DATA_BLOCK "PanelCompBAJA MTA"   // DB74
{ S7_Optimized_Access := 'FALSE' }
VERSION : 0.1
   VAR
      InhMC060 : Bool;
      InhMC061 : Bool;
      InhMC062 : Bool;
      InhMC063 : Bool;
      InhMC064 : Bool;
      InhMC065 : Bool;
      Flanco1MC060 : Bool;
      Flanco1MC061 : Bool;
      Flanco1MC062 : Bool;
      Flanco1MC063 : Bool;
      Flanco1MC064 : Bool;
      Flanco1MC065 : Bool;
      Flanco2MC060 : Bool;
      Flanco2MC061 : Bool;
      Flanco2MC062 : Bool;
      Flanco2MC063 : Bool;
      Flanco2MC064 : Bool;
      Flanco2MC065 : Bool;
      Flanco3MC060 : Bool;
      Flanco3MC061 : Bool;
      Flanco3MC062 : Bool;
      Flanco3MC063 : Bool;
      Flanco3MC064 : Bool;
      Flanco3MC065 : Bool;
      HabPanelMC060 : Bool;
      HabPanelMC061 : Bool;
      HabPanelMC062 : Bool;
      HabPanelMC063 : Bool;
      HabPanelMC064 : Bool;
      HabPanelMC065 : Bool;
      DeshabPanelMC060 : Bool;
      DeshabPanelMC061 : Bool;
      DeshabPanelMC062 : Bool;
      DeshabPanelMC063 : Bool;
      DeshabPanelMC064 : Bool;
      DeshabPanelMC065 : Bool;
      MarchaPanelMC060 : Bool;
      MarchaPanelMC061 : Bool;
      MarchaPanelMC062 : Bool;
      MarchaPanelMC063 : Bool;
      MarchaPanelMC064 : Bool;
      MarchaPanelMC065 : Bool;
      ParadaPanelMC060 : Bool;
      ParadaPanelMC061 : Bool;
      ParadaPanelMC062 : Bool;
      ParadaPanelMC063 : Bool;
      ParadaPanelMC064 : Bool;
      ParadaPanelMC065 : Bool;
      HabMC060 : Bool;
      HabMC061 : Bool;
      HabMC062 : Bool;
      HabMC063 : Bool;
      HabMC064 : Bool;
      HabMC065 : Bool;
      DeshabMC060 : Bool;
      DeshabMC061 : Bool;
      DeshabMC062 : Bool;
      DeshabMC063 : Bool;
      DeshabMC064 : Bool;
      DeshabMC065 : Bool;
      MarchaMC060 : Bool;
      MarchaMC061 : Bool;
      MarchaMC062 : Bool;
      MarchaMC063 : Bool;
      MarchaMC064 : Bool;
      MarchaMC065 : Bool;
      ParadaMC060 : Bool;
      ParadaMC061 : Bool;
      ParadaMC062 : Bool;
      ParadaMC063 : Bool;
      ParadaMC064 : Bool;
      ParadaMC065 : Bool;
      AnimMC060 : Byte;
      AnimMC061 : Byte;
      AnimMC062 : Byte;
      AnimMC063 : Byte;
      AnimMC064 : Byte;
      AnimMC065 : Byte;
      FallaGMTMC060 : Bool;
      FallaGMTMC061 : Bool;
      FallaGMTMC062 : Bool;
      FallaGMTMC063 : Bool;
      FallaGMTMC064 : Bool;
      FallaGMTMC065 : Bool;
      FallaCTCMC060 : Bool;
      FallaCTCMC061 : Bool;
      FallaCTCMC062 : Bool;
      FallaCTCMC063 : Bool;
      FallaCTCMC064 : Bool;
      FallaCTCMC065 : Bool;
      MantMC060 : Bool;
      MantMC061 : Bool;
      MantMC062 : Bool;
      MantMC063 : Bool;
      MantMC064 : Bool;
      MantMC065 : Bool;
      Reserva_1 : Bool;
      Reserva_11 : Bool;
      Reserva_12 : Bool;
      Reserva_13 : Bool;
      Reserva_14 : Bool;
      Reserva_15 : Bool;
      Reserva_16 : Bool;
      Reserva_17 : Bool;
      Reserva_18 : Bool;
      Reserva_19 : Bool;
      Reserva_110 : Bool;
      Reserva_111 : Bool;
      Reserva_112 : Bool;
      Reserva_113 : Bool;
      Reserva_114 : Bool;
      Reserva_115 : Bool;
      Reserva_116 : Bool;
      Reserva_117 : Bool;
      Reserva_118 : Bool;
      Reserva_119 : Bool;
      Reserva_120 : Bool;
      Reserva_121 : Bool;
      Reserva_122 : Bool;
      Reserva_123 : Bool;
      Reserva_124 : Bool;
      Reserva_125 : Bool;
      Reserva_126 : Bool;
      Reserva_127 : Bool;
      Reserva_128 : Bool;
      Reserva_129 : Bool;
      Reserva_130 : Bool;
      Reserva_131 : Bool;
      Reserva_132 : Bool;
      Reserva_133 : Bool;
      Reserva_134 : Bool;
      Reserva_135 : Bool;
      Reserva_136 : Bool;
      Reserva_137 : Bool;
      Reserva_138 : Bool;
      Reserva_139 : Bool;
      Reserva_140 : Bool;
      Reserva_141 : Bool;
      Reserva_142 : Bool;
      Reserva_143 : Bool;
   END_VAR
BEGIN
END_DATA_BLOCK

DATA_BLOCK "CmpBajaAuto"   // DB93
{ S7_Optimized_Access := 'FALSE' }
VERSION : 0.1
   VAR
      AutoMC060 : Bool;
      AutoMC061 : Bool;
      AutoMC062 : Bool;
      AutoMC063 : Bool;
      AutoMC064 : Bool;
      SPonMC060 : Real;
      SPonMC061 : Real;
      SPonMC062 : Real;
      SPonMC063 : Real;
      SPonMC064 : Real;
      SPoffMC060 : Real;
      SPoffMC061 : Real;
      SPoffMC062 : Real;
      SPoffMC063 : Real;
      SPoffMC064 : Real;
      AutoArrMC060 : Bool;
      AutoArrMC061 : Bool;
      AutoArrMC062 : Bool;
      AutoArrMC063 : Bool;
      AutoArrMC064 : Bool;
      AutoArrEfMC060 : Bool;
      AutoArrEfMC061 : Bool;
      AutoArrEfMC062 : Bool;
      AutoArrEfMC063 : Bool;
      AutoArrEfMC064 : Bool;
      MenuMC060 : Int;
      MenuMC061 : Int;
      MenuMC062 : Int;
      MenuMC063 : Int;
      MenuMC064 : Int;
   END_VAR
BEGIN
END_DATA_BLOCK

// folder: Entradas Analógicas

DATA_BLOCK "CaudalPotencia"   // DB26
{ S7_Optimized_Access := 'FALSE' }
VERSION : 0.1
   VAR
      lecCaudal : Real;
      lecPotencia : Real;
      HI_caudal : Real;
      LO_caudal : Real;
      HI_potencia : Real;
      LO_potencia : Real;
   END_VAR
BEGIN
END_DATA_BLOCK

DATA_BLOCK "LectAnalógicasMTA"   // DB52
{ S7_Optimized_Access := 'FALSE' }
VERSION : 0.1
   VAR
      TempCav : Real;
      TempChill : Real;
      PresAlta1 : Real;
      PresAlta12 : Real;
      PresBaja : Real;
      PreAltaHH : Real;
      PreAltaH : Real;
      PreAltaL : Real;
      PreAltaLL : Real;
      PreBajaHH : Real;
      PreBajaH : Real;
      PreBajaL : Real;
      PreBajaLL : Real;
      PresionALTA : Real;
   END_VAR
BEGIN
END_DATA_BLOCK

DATA_BLOCK "EntradasAnalógicas MTA"   // DB72
{ S7_Optimized_Access := 'FALSE' }
VERSION : 0.1
   VAR
      PresAire : Real;
      TempTanque1CH : Real;
      TempTanque2CH : Real;
      TempTorresCH : Real;
      FallaAIRE : Bool;
      FallaTanque1 : Bool;
      FallaTanque2 : Bool;
      FallaTorres : Bool;
   END_VAR
BEGIN
END_DATA_BLOCK

// folder: Horas de Marcha

DATA_BLOCK "Varios"   // DB2
{ S7_Optimized_Access := 'FALSE' }
VERSION : 0.1
   VAR
      HorasMantMC001_1 : DInt;
      HorasMantMC002_1 : DInt;
      HorasMantMC003_1 : DInt;
      HorasMantMC004_1 : DInt;
      HorasMantMC005_1 : DInt;
      HorasMantMC006_1 : DInt;
      HorasMantMC001_2 : DInt;
      HorasMantMC002_2 : DInt;
      HorasMantMC003_2 : DInt;
      HorasMantMC004_2 : DInt;
      HorasMantMC005_2 : DInt;
      HorasMantMC006_2 : DInt;
      UltimoMantMC001_1 : DInt;
      UltimoMantMC002_1 : DInt;
      UltimoMantMC003_1 : DInt;
      UltimoMantMC004_1 : DInt;
      UltimoMantMC005_1 : DInt;
      UltimoMantMC006_1 : DInt;
      UltimoMantMC001_2 : DInt;
      UltimoMantMC002_2 : DInt;
      UltimoMantMC003_2 : DInt;
      UltimoMantMC004_2 : DInt;
      UltimoMantMC005_2 : DInt;
      UltimoMantMC006_2 : DInt;
      HorasMantMS050 : DInt;
      HorasMantMS051 : DInt;
      HorasMantMS052 : DInt;
      HorasMantMS053 : DInt;
      UltimoMantMS050 : DInt;
      UltimoMantMS051 : DInt;
      UltimoMantMS052 : DInt;
      UltimoMantMS053 : DInt;
      HorasMantMC060_1 : DInt;
      HorasMantMC061_1 : DInt;
      HorasMantMC062_1 : DInt;
      HorasMantMC063_1 : DInt;
      HorasMantMC064_1 : DInt;
      HorasMantMC065_1 : DInt;
      HorasMantMC060_2 : DInt;
      HorasMantMC061_2 : DInt;
      HorasMantMC062_2 : DInt;
      HorasMantMC063_2 : DInt;
      HorasMantMC064_2 : DInt;
      HorasMantMC065_2 : DInt;
      HorasMantMC060_3 : DInt;
      HorasMantMC061_3 : DInt;
      HorasMantMC062_3 : DInt;
      HorasMantMC063_3 : DInt;
      HorasMantMC064_3 : DInt;
      HorasMantMC065_3 : DInt;
      HorasMantMC060_4 : DInt;
      HorasMantMC061_4 : DInt;
      HorasMantMC062_4 : DInt;
      HorasMantMC063_4 : DInt;
      HorasMantMC064_4 : DInt;
      HorasMantMC065_4 : DInt;
      HorasMantMC060_5 : DInt;
      HorasMantMC061_5 : DInt;
      HorasMantMC062_5 : DInt;
      HorasMantMC063_5 : DInt;
      HorasMantMC064_5 : DInt;
      HorasMantMC065_5 : DInt;
      UltimoMantMC060_1 : DInt;
      UltimoMantMC061_1 : DInt;
      UltimoMantMC062_1 : DInt;
      UltimoMantMC063_1 : DInt;
      UltimoMantMC064_1 : DInt;
      UltimoMantMC065_1 : DInt;
      UltimoMantMC060_2 : DInt;
      UltimoMantMC061_2 : DInt;
      UltimoMantMC062_2 : DInt;
      UltimoMantMC063_2 : DInt;
      UltimoMantMC064_2 : DInt;
      UltimoMantMC065_2 : DInt;
      UltimoMantMC060_3 : DInt;
      UltimoMantMC061_3 : DInt;
      UltimoMantMC062_3 : DInt;
      UltimoMantMC063_3 : DInt;
      UltimoMantMC064_3 : DInt;
      UltimoMantMC065_3 : DInt;
      UltimoMantMC060_4 : DInt;
      UltimoMantMC061_4 : DInt;
      UltimoMantMC062_4 : DInt;
      UltimoMantMC063_4 : DInt;
      UltimoMantMC064_4 : DInt;
      UltimoMantMC065_4 : DInt;
      UltimoMantMC060_5 : DInt;
      UltimoMantMC061_5 : DInt;
      UltimoMantMC062_5 : DInt;
      UltimoMantMC063_5 : DInt;
      UltimoMantMC064_5 : DInt;
      UltimoMantMC065_5 : DInt;
      HorasMantMS054_1 : DInt;
      HorasMantMS055_1 : DInt;
      HorasMantMS056_1 : DInt;
      HorasMantMS054_2 : DInt;
      HorasMantMS055_2 : DInt;
      HorasMantMS056_2 : DInt;
      UltimoMantMS054_1 : DInt;
      UltimoMantMS055_1 : DInt;
      UltimoMantMS056_1 : DInt;
      UltimoMantMS054_2 : DInt;
      UltimoMantMS055_2 : DInt;
      UltimoMantMS056_2 : DInt;
      HorasMantBost1 : DInt;
      HorasMantBost2 : DInt;
      UltimoMantBoost1 : DInt;
      UltimoMantBoost2 : DInt;
   END_VAR
BEGIN
END_DATA_BLOCK

DATA_BLOCK "HorasSecAlta"   // DB19
{ S7_Optimized_Access := 'FALSE' }
VERSION : 0.1
   VAR
      HMMS050 : DInt;
      HMMS051 : DInt;
      HMMS052 : DInt;
      HMMS053 : DInt;
      MMMS050 : Int;
      MMMS051 : Int;
      MMMS052 : Int;
      MMMS053 : Int;
      SMMS050 : Int;
      SMMS051 : Int;
      SMMS052 : Int;
      SMMS053 : Int;
   END_VAR
BEGIN
END_DATA_BLOCK

DATA_BLOCK "HorasCmpBaja"   // DB20
{ S7_Optimized_Access := 'FALSE' }
VERSION : 0.1
   VAR
      HMMC060 : DInt;
      HMMC061 : DInt;
      HMMC062 : DInt;
      HMMC063 : DInt;
      HMMC064 : DInt;
      HMMC065 : DInt;
      MMMC060 : Int;
      MMMC061 : Int;
      MMMC062 : Int;
      MMMC063 : Int;
      MMMC064 : Int;
      MMMC065 : Int;
      SMMC060 : Int;
      SMMC061 : Int;
      SMMC062 : Int;
      SMMC063 : Int;
      SMMC064 : Int;
      SMMC065 : Int;
   END_VAR
BEGIN
END_DATA_BLOCK

DATA_BLOCK "HorasSecBaja"   // DB24
{ S7_Optimized_Access := 'FALSE' }
VERSION : 0.1
   VAR
      HMMS054 : DInt;
      HMMS055 : DInt;
      HMMS056 : DInt;
      MMMS054 : Int;
      MMMS055 : Int;
      MMMS056 : Int;
      SMMS054 : Int;
      SMMS055 : Int;
      SMMS056 : Int;
   END_VAR
BEGIN
END_DATA_BLOCK

DATA_BLOCK "SumaOB35 MTA"   // DB73
{ S7_Optimized_Access := 'FALSE' }
VERSION : 0.1
   VAR
      HMMC001 : DInt;
      HMMC002 : DInt;
      HMMC003 : DInt;
      HMMC004 : DInt;
      HMMC005 : DInt;
      HMMC006 : DInt;
      MMMC001 : Int;
      MMMC002 : Int;
      MMMC003 : Int;
      MMMC004 : Int;
      MMMC005 : Int;
      MMMC006 : Int;
      PrioridadArranqueMC001 : Int;
      PrioridadArranqueMC002 : Int;
      PrioridadArranqueMC003 : Int;
      PrioridadArranqueMC004 : Int;
      PrioridadArranqueMC005 : Int;
      PrioridadArranqueMC006 : Int;
      PrioridadParadaMC001 : Int;
      PrioridadParadaMC002 : Int;
      PrioridadParadaMC003 : Int;
      PrioridadParadaMC004 : Int;
      PrioridadParadaMC005 : Int;
      PrioridadParadaMC006 : Int;
      HorasMin : DInt;
      HorasMax : DInt;
      MotoreEnMarcha : Int;
      SMMC001 : Int;
      SMMC002 : Int;
      SMMC003 : Int;
      SMMC004 : Int;
      SMMC005 : Int;
      SMMC006 : Int;
      ByteMotoresEnAUTO : Byte;
      ByteMotoresEnMarcha : Byte;
   END_VAR
BEGIN
END_DATA_BLOCK

// folder: Iluminación

DATA_BLOCK "DBIluminaciónMTA"   // DB87
{ S7_Optimized_Access := 'FALSE' }
VERSION : 0.1
   VAR
      TiempoDeEncendido : Word;
      EncendidoPanel : Bool;
      ApagadoPanel : Bool;
      Encendido : Bool;
      MantenerEncendida : Bool;
      AuxiliarEncendidoPermane : Bool;
      FLANCOP : Bool;
      FLANCON : Bool;
      EcendidoPLS : Bool;
      ApagadoPLS : Bool;
      TiempoPANEL : S5Time;
      AuxiliarCalculo : Int;
      TiempoPANEL1 : S5Time;
   END_VAR
BEGIN
END_DATA_BLOCK

// folder: Panel

DATA_BLOCK "Bloque de animacion MTA"   // DB46
{ S7_Optimized_Access := 'FALSE' }
VERSION : 0.1
   VAR
      AnimacionMP010 : Byte;
      AnimacionMP011 : Byte;
      AnimacionMP012 : Byte;
      AnimacionMP013 : Byte;
      AnimacionMP018 : Byte;
      AnimacionMP019 : Byte;
      AnimacionMT007 : Byte;
      AnimacionMT008 : Byte;
      AnimacionMT009 : Byte;
      AnimacionMT010 : Byte;
      AnimacionV001 : Byte;
      AnimacionV002 : Byte;
      AnimacionV003 : Byte;
      MenuMS050 : Int;
      MenuMS051 : Int;
      MenuMS052 : Int;
      MenuMS053 : Int;
      MenuMS054 : Int;
      MenuV001 : Int;
      MenuV002 : Int;
      MenuV003 : Int;
      AnimacionMS054 : Byte;
      AnimacionMS055 : Byte;
      MenuV030 : Int;
      MenuV031 : Int;
      AnimMV030 : Byte;
      AnimMV031 : Byte;
      AnimMP014 : Byte;
      AnimMP015 : Byte;
      AnimMC001 : Byte;
      AnimMC002 : Byte;
      AnimMC003 : Byte;
      AnimMC004 : Byte;
      AnimMC005 : Byte;
      AnimMC006 : Byte;
      Reserva17 : Byte;
      Reserva18 : Byte;
      Reserva19 : Byte;
      Reserva20 : Byte;
      Reserva21 : Byte;
      Reserva22 : Byte;
      Reserva23 : Byte;
      Reserva24 : Byte;
      Reserva25 : Byte;
      Reserva26 : Byte;
      Reserva27 : Byte;
      Reserva28 : Byte;
      Reserva29 : Byte;
      Reserva30 : Byte;
      Reserva31 : Byte;
      Reserva32 : Byte;
      Reserva33 : Byte;
      Reserva34 : Byte;
      Reserva35 : Byte;
      Reserva36 : Byte;
      Reserva37 : Byte;
      Reserva38 : Byte;
      Reserva39 : Byte;
      Reserva40 : Byte;
      Reserva41 : Byte;
      Reserva42 : Byte;
      Reserva43 : Byte;
      Reserva44 : Byte;
      Reserva45 : Byte;
      Reserva46 : Byte;
      Reserva47 : Byte;
      Reserva48 : Byte;
      Reserva49 : Byte;
      Reserva50 : Byte;
      Reserva51 : Byte;
      Reserva52 : Byte;
      Reserva53 : Byte;
      Reserva54 : Byte;
      Reserva55 : Byte;
      Reserva56 : Byte;
      Reserva57 : Byte;
      Reserva58 : Byte;
      Reserva59 : Byte;
      Reserva60 : Byte;
      Reserva61 : Byte;
      Reserva62 : Byte;
      Reserva63 : Byte;
      Reserva64 : Byte;
      Reserva65 : Byte;
      Reserva66 : Byte;
      Reserva67 : Byte;
      Reserva68 : Byte;
      Reserva69 : Byte;
      Reserva70 : Byte;
      Reserva71 : Byte;
      Reserva72 : Byte;
      Reserva73 : Byte;
      Reserva74 : Byte;
   END_VAR
BEGIN
END_DATA_BLOCK

DATA_BLOCK "PanelMotChillMTA"   // DB90
{ S7_Optimized_Access := 'FALSE' }
VERSION : 0.1
   VAR
      InhMT007 : Bool;
      InhMT008 : Bool;
      InhMT009 : Bool;
      InhMT010 : Bool;
      InhMP010 : Bool;
      InhMP011 : Bool;
      InhMP012 : Bool;
      InhMP013 : Bool;
      InhMP018 : Bool;
      InhMP019 : Bool;
      InhV001 : Bool;
      InhV002 : Bool;
      InhV003 : Bool;
      Flanco1MT007 : Bool;
      Flanco1MT008 : Bool;
      Flanco1MT009 : Bool;
      Flanco1MT010 : Bool;
      Flanco1MP010 : Bool;
      Flanco1MP011 : Bool;
      Flanco1MP012 : Bool;
      Flanco1MP013 : Bool;
      Flanco1MP018 : Bool;
      Flanco1MP019 : Bool;
      Flanco1V001 : Bool;
      Flanco1V002 : Bool;
      Flanco1V003 : Bool;
      Flanco2MT007 : Bool;
      Flanco2MT008 : Bool;
      Flanco2MT009 : Bool;
      Flanco2MT010 : Bool;
      Flanco2MP010 : Bool;
      Flanco2MP011 : Bool;
      Flanco2MP012 : Bool;
      Flanco2MP013 : Bool;
      Flanco2MP018 : Bool;
      Flanco2MP019 : Bool;
      Flanco2V001 : Bool;
      Flanco2V002 : Bool;
      Flanco2V003 : Bool;
      Flanco3MT007 : Bool;
      Flanco3MT008 : Bool;
      Flanco3MT009 : Bool;
      Flanco3MT010 : Bool;
      Flanco3MP010 : Bool;
      Flanco3MP011 : Bool;
      Flanco3MP012 : Bool;
      Flanco3MP013 : Bool;
      Flanco3MP018 : Bool;
      Flanco3MP019 : Bool;
      Flanco3V001 : Bool;
      Flanco3V002 : Bool;
      Flanco3V003 : Bool;
      HabPanelMT007 : Bool;
      HabPanelMT008 : Bool;
      HabPanelMT009 : Bool;
      HabPanelMT010 : Bool;
      HabPanelMP010 : Bool;
      HabPanelMP011 : Bool;
      HabPanelMP012 : Bool;
      HabPanelMP013 : Bool;
      HabPanelMP018 : Bool;
      HabPanelMP019 : Bool;
      HabPanelV001 : Bool;
      HabPanelV002 : Bool;
      HabPanelV003 : Bool;
      DeshabPanelMT007 : Bool;
      DeshabPanelMT008 : Bool;
      DeshabPanelMT009 : Bool;
      DeshabPanelMT010 : Bool;
      DeshabPanelMP010 : Bool;
      DeshabPanelMP011 : Bool;
      DeshabPanelMP012 : Bool;
      DeshabPanelMP013 : Bool;
      DeshabPanelMP018 : Bool;
      DeshabPanelMP019 : Bool;
      DeshabPanelV001 : Bool;
      DeshabPanelV002 : Bool;
      DeshabPanelV003 : Bool;
      MarchaPanelMT007 : Bool;
      MarchaPanelMT008 : Bool;
      MarchaPanelMT009 : Bool;
      MarchaPanelMT010 : Bool;
      MarchaPanelMP010 : Bool;
      MarchaPanelMP011 : Bool;
      MarchaPanelMP012 : Bool;
      MarchaPanelMP013 : Bool;
      MarchaPanelMP018 : Bool;
      MarchaPanelMP019 : Bool;
      MarchaPanelV001 : Bool;
      MarchaPanelV002 : Bool;
      MarchaPanelV003 : Bool;
      ParadaPanelMT007 : Bool;
      ParadaPanelMT008 : Bool;
      ParadaPanelMT009 : Bool;
      ParadaPanelMT010 : Bool;
      ParadaPanelMP010 : Bool;
      ParadaPanelMP011 : Bool;
      ParadaPanelMP012 : Bool;
      ParadaPanelMP013 : Bool;
      ParadaPanelMP018 : Bool;
      ParadaPanelMP019 : Bool;
      ParadaPanelV001 : Bool;
      ParadaPanelV002 : Bool;
      ParadaPanelV003 : Bool;
      HabMT007 : Bool;
      HabMT008 : Bool;
      HabMT009 : Bool;
      HabMT010 : Bool;
      HabMP010 : Bool;
      HabMP011 : Bool;
      HabMP012 : Bool;
      HabMP013 : Bool;
      HabMP018 : Bool;
      HabMP019 : Bool;
      HabV001 : Bool;
      HabV002 : Bool;
      HabV003 : Bool;
      DeshabMT007 : Bool;
      DeshabMT008 : Bool;
      DeshabMT009 : Bool;
      DeshabMT010 : Bool;
      DeshabMP010 : Bool;
      DeshabMP011 : Bool;
      DeshabMP012 : Bool;
      DeshabMP013 : Bool;
      DeshabMP018 : Bool;
      DeshabMP019 : Bool;
      DeshabV001 : Bool;
      DeshabV002 : Bool;
      DeshabV003 : Bool;
      MarchaMT007 : Bool;
      MarchaMT008 : Bool;
      MarchaMT009 : Bool;
      MarchaMT010 : Bool;
      MarchaMP010 : Bool;
      MarchaMP011 : Bool;
      MarchaMP012 : Bool;
      MarchaMP013 : Bool;
      MarchaMP018 : Bool;
      MarchaMP019 : Bool;
      MarchaV001 : Bool;
      MarchaV002 : Bool;
      MarchaV003 : Bool;
      ParadaMT007 : Bool;
      ParadaMT008 : Bool;
      ParadaMT009 : Bool;
      ParadaMT010 : Bool;
      ParadaMP010 : Bool;
      ParadaMP011 : Bool;
      ParadaMP012 : Bool;
      ParadaMP013 : Bool;
      ParadaMP018 : Bool;
      ParadaMP019 : Bool;
      ParadaV001 : Bool;
      ParadaV002 : Bool;
      ParadaV003 : Bool;
      AnimMT007 : Byte;
      AnimMT008 : Byte;
      AnimMT009 : Byte;
      AnimMT010 : Byte;
      AnimMP010 : Byte;
      AnimMP011 : Byte;
      AnimMP012 : Byte;
      AnimMP013 : Byte;
      AnimMP018 : Byte;
      AnimMP019 : Byte;
      AnimV001 : Byte;
      AnimV002 : Byte;
      AnimV003 : Byte;
      Reserva_1 : Bool;
      Reserva_11 : Bool;
      Reserva_12 : Bool;
      Reserva_13 : Bool;
      Reserva_14 : Bool;
      Reserva_15 : Bool;
      Reserva_16 : Bool;
      Reserva_17 : Bool;
      Reserva_18 : Bool;
      Reserva_19 : Bool;
      Reserva_110 : Bool;
      Reserva_111 : Bool;
      Reserva_112 : Bool;
      Reserva_113 : Bool;
      Reserva_114 : Bool;
      Reserva_115 : Bool;
      Reserva_116 : Bool;
      Reserva_117 : Bool;
      Reserva_118 : Bool;
      Reserva_119 : Bool;
      Reserva_120 : Bool;
      Reserva_121 : Bool;
      Reserva_122 : Bool;
      Reserva_123 : Bool;
      Reserva_124 : Bool;
      Reserva_125 : Bool;
      Reserva_126 : Bool;
      Reserva_127 : Bool;
      Reserva_128 : Bool;
      Reserva_129 : Bool;
      Reserva_130 : Bool;
      Reserva_131 : Bool;
      Reserva_132 : Bool;
      Reserva_133 : Bool;
      Reserva_134 : Bool;
      Reserva_135 : Bool;
      Reserva_136 : Bool;
      Reserva_137 : Bool;
      Reserva_138 : Bool;
      Reserva_139 : Bool;
      Reserva_140 : Bool;
      Reserva_141 : Bool;
      Reserva_142 : Bool;
      Reserva_143 : Bool;
   END_VAR
BEGIN
END_DATA_BLOCK

// folder: Secadores/Alta

DATA_BLOCK "PanelSecALTA"   // DB81
{ S7_Optimized_Access := 'FALSE' }
VERSION : 0.1
   VAR
      InhMS050 : Bool;
      InhMS051 : Bool;
      InhMS052 : Bool;
      InhMS053 : Bool;
      Flanco1MS050 : Bool;
      Flanco1MS051 : Bool;
      Flanco1MS052 : Bool;
      Flanco1MS053 : Bool;
      Flanco2MS050 : Bool;
      Flanco2MS051 : Bool;
      Flanco2MS052 : Bool;
      Flanco2MS053 : Bool;
      Flanco3MS050 : Bool;
      Flanco3MS051 : Bool;
      Flanco3MS052 : Bool;
      Flanco3MS053 : Bool;
      HabPanelMS050 : Bool;
      HabPanelMS051 : Bool;
      HabPanelMS052 : Bool;
      HabPanelMS053 : Bool;
      DeshabPanelMS050 : Bool;
      DeshabPanelMS051 : Bool;
      DeshabPanelMS052 : Bool;
      DeshabPanelMS053 : Bool;
      MarchaPanelMS050 : Bool;
      MarchaPanelMS051 : Bool;
      MarchaPanelMS052 : Bool;
      MarchaPanelMS053 : Bool;
      ParadaPanelMS050 : Bool;
      ParadaPanelMS051 : Bool;
      ParadaPanelMS052 : Bool;
      ParadaPanelMS053 : Bool;
      HabMS050 : Bool;
      HabMS051 : Bool;
      HabMS052 : Bool;
      HabMS053 : Bool;
      DeshabMS050 : Bool;
      DeshabMS051 : Bool;
      DeshabMS052 : Bool;
      DeshabMS053 : Bool;
      MarchaMS050 : Bool;
      MarchaMS051 : Bool;
      MarchaMS052 : Bool;
      MarchaMS053 : Bool;
      ParadaMS050 : Bool;
      ParadaMS051 : Bool;
      ParadaMS052 : Bool;
      ParadaMS053 : Bool;
      AnimMS050 : Byte;
      AnimMS051 : Byte;
      AnimMS052 : Byte;
      AnimMS053 : Byte;
      FallaGMTMS050 : Bool;
      FallaGMTMS051 : Bool;
      FallaGMTMS052 : Bool;
      FallaGMTMS053 : Bool;
      FallaCTCMS050 : Bool;
      FallaCTCMS051 : Bool;
      FallaCTCMS052 : Bool;
      FallaCTCMS053 : Bool;
      MantMS050 : Bool;
      MantMS051 : Bool;
      MantMS052 : Bool;
      MantMS053 : Bool;
      Enc1MS050 : Int;
      Enc2MS050 : Int;
      Enc1MS051 : Int;
      Enc2MS051 : Int;
      Enc1MS052 : Int;
      Enc2MS052 : Int;
      Enc1MS053 : Int;
      Enc2MS053 : Int;
      AutoMS050 : Bool;
      AutoMS051 : Bool;
      AutoMS052 : Bool;
      AutoMS053 : Bool;
      AutoArrMS050 : Bool;
      AutoArrMS051 : Bool;
      AutoArrMS052 : Bool;
      AutoArrMS053 : Bool;
      Reserva2 : Bool;
      Reserva3 : Bool;
      Reserva4 : Bool;
      Reserva_15 : Bool;
      Reserva_16 : Bool;
      Reserva_17 : Bool;
      Reserva_18 : Bool;
      Reserva_19 : Bool;
      Reserva_110 : Bool;
      Reserva_111 : Bool;
      Reserva_112 : Bool;
      Reserva_113 : Bool;
      Reserva_114 : Bool;
      Reserva_115 : Bool;
      Reserva_116 : Bool;
      Reserva_117 : Bool;
      Reserva_118 : Bool;
      Reserva_119 : Bool;
      Reserva_120 : Bool;
      Reserva_121 : Bool;
      Reserva_122 : Bool;
      Reserva_123 : Bool;
      Reserva_124 : Bool;
      Reserva_125 : Bool;
      Reserva_126 : Bool;
      Reserva_127 : Bool;
      Reserva_128 : Bool;
      Reserva_129 : Bool;
      Reserva_130 : Bool;
      Reserva_131 : Bool;
      Reserva_132 : Bool;
      Reserva_133 : Bool;
      Reserva_134 : Bool;
      Reserva_135 : Bool;
      Reserva_136 : Bool;
      Reserva_137 : Bool;
      Reserva_138 : Bool;
      Reserva_139 : Bool;
      Reserva_140 : Bool;
      Reserva_141 : Bool;
      Reserva_142 : Bool;
      Reserva_143 : Bool;
   END_VAR
BEGIN
END_DATA_BLOCK

// folder: Secadores/Baja

DATA_BLOCK "PanelSecBaja"   // DB49
{ S7_Optimized_Access := 'FALSE' }
VERSION : 0.1
   VAR
      InhMS054 : Bool;
      InhMS055 : Bool;
      Flanco1MS054 : Bool;
      Flanco1MS055 : Bool;
      Flanco2MS054 : Bool;
      Flanco2MS055 : Bool;
      Flanco3MS054 : Bool;
      Flanco3MS055 : Bool;
      HabPanelMS054 : Bool;
      HabPanelMS055 : Bool;
      DeshabPanelMS054 : Bool;
      DeshabPanelMS055 : Bool;
      MarchaPanelMS054 : Bool;
      MarchaPanelMS055 : Bool;
      ParadaPanelMS054 : Bool;
      ParadaPanelMS055 : Bool;
      HabMS054 : Bool;
      HabMS055 : Bool;
      DeshabMS054 : Bool;
      DeshabMS055 : Bool;
      MarchaMS054 : Bool;
      MarchaMS055 : Bool;
      ParadaMS054 : Bool;
      ParadaMS055 : Bool;
      AnimMS054 : Byte;
      AnimMS055 : Byte;
      FallaGMTMS054 : Bool;
      FallaGMTMS055 : Bool;
      FallaCTCMS054 : Bool;
      FallaCTCMS055 : Bool;
      MantMS054 : Bool;
      MantMS055 : Bool;
      Reserva2 : Bool;
      Reserva3 : Bool;
      Reserva4 : Bool;
      Reserva_15 : Bool;
      Reserva_16 : Bool;
      Reserva_17 : Bool;
      Reserva_18 : Bool;
      Reserva_19 : Bool;
      Reserva_110 : Bool;
      Reserva_111 : Bool;
      Reserva_112 : Bool;
      Reserva_113 : Bool;
      Reserva_114 : Bool;
      Reserva_115 : Bool;
      Reserva_116 : Bool;
      Reserva_117 : Bool;
      Reserva_118 : Bool;
      Reserva_119 : Bool;
      Reserva_120 : Bool;
      Reserva_121 : Bool;
      Reserva_122 : Bool;
      Reserva_123 : Bool;
      Reserva_124 : Bool;
      Reserva_125 : Bool;
      Reserva_126 : Bool;
      Reserva_127 : Bool;
      Reserva_128 : Bool;
      Reserva_129 : Bool;
      Reserva_130 : Bool;
      Reserva_131 : Bool;
      Reserva_132 : Bool;
      Reserva_133 : Bool;
      Reserva_134 : Bool;
      Reserva_135 : Bool;
      Reserva_136 : Bool;
      Reserva_137 : Bool;
      Reserva_138 : Bool;
      Reserva_139 : Bool;
      Reserva_140 : Bool;
      Reserva_141 : Bool;
      Reserva_142 : Bool;
      Reserva_143 : Bool;
   END_VAR
BEGIN
END_DATA_BLOCK

// folder: Torres de Agua/Torres Cavaleto

DATA_BLOCK "PanelTorreCav"   // DB21
{ S7_Optimized_Access := 'FALSE' }
VERSION : 0.1
   VAR
      InhMV030 : Bool;
      InhMV031 : Bool;
      InhMP014 : Bool;
      InhMP015 : Bool;
      Flanco1MV030 : Bool;
      Flanco1MV031 : Bool;
      Flanco1MP014 : Bool;
      Flanco1MP015 : Bool;
      Flanco2MV030 : Bool;
      Flanco2MV031 : Bool;
      Flanco2MP014 : Bool;
      Flanco2MP015 : Bool;
      Flanco3MV030 : Bool;
      Flanco3MV031 : Bool;
      Flanco3MP014 : Bool;
      Flanco3MP015 : Bool;
      HabPanelMV030 : Bool;
      HabPanelMV031 : Bool;
      HabPanelMP014 : Bool;
      HabPanelMP015 : Bool;
      DeshabPanelMV030 : Bool;
      DeshabPanelMV031 : Bool;
      DeshabPanelMP014 : Bool;
      DeshabPanelMP015 : Bool;
      MarchaPanelMV030 : Bool;
      MarchaPanelMV031 : Bool;
      MarchaPanelMP014 : Bool;
      MarchaPanelMP015 : Bool;
      ParadaPanelMV030 : Bool;
      ParadaPanelMV031 : Bool;
      ParadaPanelMP014 : Bool;
      ParadaPanelMP015 : Bool;
      HabMV030 : Bool;
      HabMV031 : Bool;
      HabMP014 : Bool;
      HabMP015 : Bool;
      DeshabMV030 : Bool;
      DeshabMV031 : Bool;
      DeshabMP014 : Bool;
      DeshabMP015 : Bool;
      MarchaMV030 : Bool;
      MarchaMV031 : Bool;
      MarchaMP014 : Bool;
      MarchaMP015 : Bool;
      ParadaMV030 : Bool;
      ParadaMV031 : Bool;
      ParadaMP014 : Bool;
      ParadaMP015 : Bool;
      MantMV030 : Bool;
      MantMV031 : Bool;
      MantMP014 : Bool;
      MantMP015 : Bool;
      AutoV030 : Bool;
      AutoV031 : Bool;
      SPonV030 : Int;
      SPonV031 : Int;
      SPoffV030 : Int;
      SPoffV031 : Int;
      Temperatura : Int;
      ArranqueAutoV030 : Bool;
      ArranqueAutoV031 : Bool;
      Reserva_13 : Bool;
      Reserva_14 : Bool;
      Reserva_15 : Bool;
      Reserva_16 : Bool;
      Reserva_17 : Bool;
      Reserva_18 : Bool;
      Reserva_19 : Bool;
      Reserva_110 : Bool;
      Reserva_111 : Bool;
      Reserva_112 : Bool;
      Reserva_113 : Bool;
      Reserva_114 : Bool;
      Reserva_115 : Bool;
      Reserva_116 : Bool;
      Reserva_117 : Bool;
      Reserva_118 : Bool;
      Reserva_119 : Bool;
      Reserva_120 : Bool;
      Reserva_121 : Bool;
      Reserva_122 : Bool;
      Reserva_123 : Bool;
      Reserva_124 : Bool;
      Reserva_125 : Bool;
      Reserva_126 : Bool;
      Reserva_127 : Bool;
      Reserva_128 : Bool;
      Reserva_129 : Bool;
      Reserva_130 : Bool;
      Reserva_131 : Bool;
      Reserva_132 : Bool;
      Reserva_133 : Bool;
      Reserva_134 : Bool;
      Reserva_135 : Bool;
      Reserva_136 : Bool;
      Reserva_137 : Bool;
      Reserva_138 : Bool;
      Reserva_139 : Bool;
      Reserva_140 : Bool;
      Reserva_141 : Bool;
      Reserva_142 : Bool;
      Reserva_143 : Bool;
   END_VAR
BEGIN
END_DATA_BLOCK

DATA_BLOCK "TAguaCAV"   // DB51
{ S7_Optimized_Access := 'FALSE' }
AUTHOR : AEB
VERSION : 0.1
   VAR
      PrAlta : Real;
      TmpCav : Real;
      PrAlta2 : Real;
      PrBaja : Real;
      STAT4 : Real;
      STAT5 : Real;
      STAT6 : Real;
      STAT7 : Real;
      STAT8 : Real;
      STAT9 : Real;
      STAT10 : Real;
      STAT11 : Real;
      STAT12 : Real;
      STAT13 : Real;
      STAT14 : Real;
      STAT15 : Real;
      STAT16 : Real;
      STAT17 : Real;
      STAT18 : Real;
      STAT19 : Real;
      STAT20 : Real;
      STAT21 : Real;
      STAT22 : Real;
      STAT23 : Real;
      STAT24 : Real;
      STAT25 : Real;
      STAT26 : Real;
      STAT27 : Real;
      STAT28 : Real;
      STAT29 : Real;
      STAT30 : Real;
      STAT31 : Real;
      STAT32 : Real;
      STAT33 : Real;
      STAT34 : Real;
      STAT35 : Real;
      STAT36 : Real;
      STAT37 : Real;
      STAT38 : Real;
      STAT39 : Real;
      STAT40 : Real;
      STAT41 : Real;
      STAT42 : Real;
      STAT43 : Real;
      STAT44 : Real;
      STAT45 : Real;
      STAT46 : Real;
      STAT47 : Real;
      STAT48 : Real;
      STAT49 : Real;
      STAT50 : Real;
      STAT51 : Real;
      STAT52 : Real;
      STAT53 : Real;
      STAT54 : Real;
      STAT55 : Real;
      STAT56 : Real;
      STAT57 : Real;
      STAT58 : Real;
      STAT59 : Real;
      STAT60 : Real;
      STAT61 : Real;
      STAT62 : Real;
      STAT63 : Real;
      STAT64 : Real;
      STAT65 : Real;
   END_VAR
BEGIN
END_DATA_BLOCK

// folder: Torres de Agua/Torres Chillers

DATA_BLOCK "CFG-TorresCH"   // DB92
{ S7_Optimized_Access := 'FALSE' }
VERSION : 0.1
   VAR
      AutoV001 : Bool;
      AutoV002 : Bool;
      AutoV003 : Bool;
      SPonV001 : Int;
      SPonV002 : Int;
      SPonV003 : Int;
      SPoffV001 : Int;
      SPoffV002 : Int;
      SPoffV003 : Int;
      Temperatura : Int;
      ArranqueAutoV001 : Bool;
      ArranqueAutoV002 : Bool;
      ArranqueAutoV003 : Bool;
   END_VAR
BEGIN
END_DATA_BLOCK

// folder: (top level)

FUNCTION "Arranques General" : Void   // FC4, LAD
{ S7_Optimized_Access := 'FALSE' }
VERSION : 0.1
   VAR_TEMP   // added for the SCL form of the ladder/FBD networks
      _w1 : Bool;
      _w2 : Bool;
      _s5time1 : S5Time;
   END_VAR
BEGIN

REGION Network 1: Motor MT007 / Bloque motor MT007 - Bomba Soplado L1
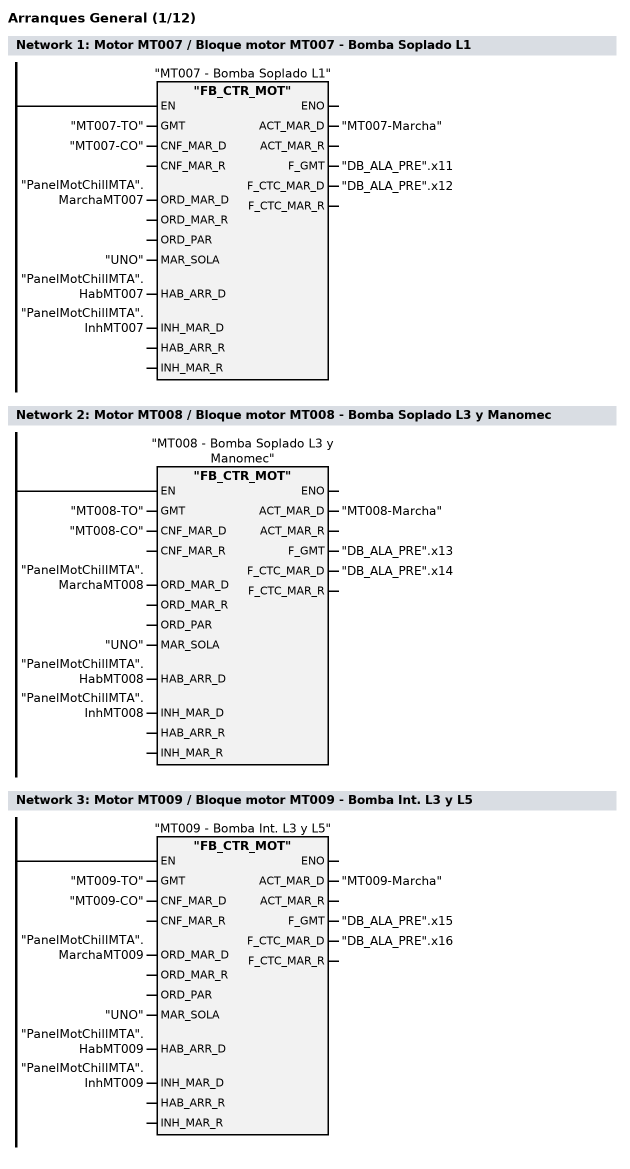
   RUNG wire#powerrail
      "MT007 - Bomba Soplado L1"(GMT := "MT007-TO", CNF_MAR_D := "MT007-CO", CNF_MAR_R :=, ORD_MAR_D := "PanelMotChillMTA".MarchaMT007, ORD_MAR_R :=, ORD_PAR :=, MAR_SOLA := "UNO", HAB_ARR_D := "PanelMotChillMTA".HabMT007, INH_MAR_D := "PanelMotChillMTA".InhMT007, HAB_ARR_R :=, INH_MAR_R :=, ACT_MAR_D => "MT007-Marcha", ACT_MAR_R =>, F_GMT => "DB_ALA_PRE".x11, F_CTC_MAR_D => "DB_ALA_PRE".x12, F_CTC_MAR_R =>)
   END_RUNG
   // the same network as SCL:
   "MT007 - Bomba Soplado L1"(GMT := "MT007-TO",   // "FB_CTR_MOT"
                           CNF_MAR_D := "MT007-CO",
                           ORD_MAR_D := "PanelMotChillMTA".MarchaMT007,
                           MAR_SOLA := "UNO",
                           HAB_ARR_D := "PanelMotChillMTA".HabMT007,
                           INH_MAR_D := "PanelMotChillMTA".InhMT007,
                           ACT_MAR_D => "MT007-Marcha",
                           F_GMT => "DB_ALA_PRE".x11,
                           F_CTC_MAR_D => "DB_ALA_PRE".x12);
END_REGION

REGION Network 2: Motor MT008 / Bloque motor MT008 - Bomba Soplado L3 y Manomec
   RUNG wire#powerrail
      "MT008 - Bomba Soplado L3 y Manomec"(GMT := "MT008-TO", CNF_MAR_D := "MT008-CO", CNF_MAR_R :=, ORD_MAR_D := "PanelMotChillMTA".MarchaMT008, ORD_MAR_R :=, ORD_PAR :=, MAR_SOLA := "UNO", HAB_ARR_D := "PanelMotChillMTA".HabMT008, INH_MAR_D := "PanelMotChillMTA".InhMT008, HAB_ARR_R :=, INH_MAR_R :=, ACT_MAR_D => "MT008-Marcha", ACT_MAR_R =>, F_GMT => "DB_ALA_PRE".x13, F_CTC_MAR_D => "DB_ALA_PRE".x14, F_CTC_MAR_R =>)
   END_RUNG
   // the same network as SCL:
   "MT008 - Bomba Soplado L3 y Manomec"(GMT := "MT008-TO",   // "FB_CTR_MOT"
                           CNF_MAR_D := "MT008-CO",
                           ORD_MAR_D := "PanelMotChillMTA".MarchaMT008,
                           MAR_SOLA := "UNO",
                           HAB_ARR_D := "PanelMotChillMTA".HabMT008,
                           INH_MAR_D := "PanelMotChillMTA".InhMT008,
                           ACT_MAR_D => "MT008-Marcha",
                           F_GMT => "DB_ALA_PRE".x13,
                           F_CTC_MAR_D => "DB_ALA_PRE".x14);
END_REGION

REGION Network 3: Motor MT009 / Bloque motor MT009 - Bomba Int. L3 y L5
   RUNG wire#powerrail
      "MT009 - Bomba Int. L3 y L5"(GMT := "MT009-TO", CNF_MAR_D := "MT009-CO", CNF_MAR_R :=, ORD_MAR_D := "PanelMotChillMTA".MarchaMT009, ORD_MAR_R :=, ORD_PAR :=, MAR_SOLA := "UNO", HAB_ARR_D := "PanelMotChillMTA".HabMT009, INH_MAR_D := "PanelMotChillMTA".InhMT009, HAB_ARR_R :=, INH_MAR_R :=, ACT_MAR_D => "MT009-Marcha", ACT_MAR_R =>, F_GMT => "DB_ALA_PRE".x15, F_CTC_MAR_D => "DB_ALA_PRE".x16, F_CTC_MAR_R =>)
   END_RUNG
   // the same network as SCL:
   "MT009 - Bomba Int. L3 y L5"(GMT := "MT009-TO",   // "FB_CTR_MOT"
                           CNF_MAR_D := "MT009-CO",
                           ORD_MAR_D := "PanelMotChillMTA".MarchaMT009,
                           MAR_SOLA := "UNO",
                           HAB_ARR_D := "PanelMotChillMTA".HabMT009,
                           INH_MAR_D := "PanelMotChillMTA".InhMT009,
                           ACT_MAR_D => "MT009-Marcha",
                           F_GMT => "DB_ALA_PRE".x15,
                           F_CTC_MAR_D => "DB_ALA_PRE".x16);
END_REGION

REGION Network 4: Motor MT010 / Bloque motor MT010 - Bomba Int L1 y Manomec